// TIA Portal project "ModBus_Tcp_ESP32_V20" (V20)
// Modbus TCP/IP connection with ESP32 microcontroller

(* hardware
DEVICE "S7-1200 station_1"  S7-1200 Station
   slot 0: "Rack_0"  S7-1200 Rack  Rack  V1.0
   slot 1: "PLC_1"  CPU 1212C AC/DC/Rly  6ES7 212-1BE40-0XB0  V4.6
DEVICE "HMI_1"  TP700 Comfort
   slot 0: "HMI_1"  TP700 Comfort  6AV2 124-0GC01-0AX0  17.0.0.0
   slot 1: "HMI_RT_1"  TP700 Comfort  6AV2 124-0GC01-0AX0  17.0.0.0
   slot 5: "HMI_1.IE_CP_1"  PROFINET Interface  17.0.0.0
      slot 1: "PROFINET Interface_1"  PROFINET Interface
         slot 1: "Port_1"  Port
         slot 2: "Port_2"  Port
   slot 7: "HMI_1.MPI/DP_CP_1"  MPI/DP Interface  17.0.0.0
*)

// ===== PLC "PLC_1"  CPU 1212C AC/DC/Rly =====

VAR_GLOBAL   // PLC tag table "Default tag table"
   "Clock_Byte" AT %MB0 : Byte;
   "Clock_10Hz" AT %M0.0 : Bool;
   "Clock_5Hz" AT %M0.1 : Bool;
   "Clock_2.5Hz" AT %M0.2 : Bool;
   "Clock_2Hz" AT %M0.3 : Bool;
   "Clock_1.25Hz" AT %M0.4 : Bool;
   "Clock_1Hz" AT %M0.5 : Bool;
   "Clock_0.625Hz" AT %M0.6 : Bool;
   "Clock_0.5Hz" AT %M0.7 : Bool;
   "Tag_1" AT %MW1 : Word;
   "Tag_2" AT %M10.1 : Bool;
   "Tag_3" AT %M10.5 : Bool;
   "Tag_4" AT %M100.1 : Bool;
   "Tag_5" AT %M10.6 : Bool;
   "Tag_6" AT %M11.1 : Bool;
   "Tag_7" AT %M12.1 : Bool;
   "Tag_8" AT %M10.0 : Bool;
END_VAR

DATA_BLOCK "Modbus_Receiver"   // DB2
{ S7_Optimized_Access := 'FALSE' }
VERSION : 0.1
   VAR
      Receiver : Array[0..7] of Word;
      ADDR : UDInt := 400001;   // Initial Address Holding Register
      DATA_LEN : UInt := 8;   // Holding Register to Read
   END_VAR
BEGIN
   // Receiver[0] : First Address
   // Receiver[4] : Command
   // Receiver[3] : Value
   // Receiver[2] : Third Address
   // Receiver[1] : Second Address
   // Receiver[5] : Frequency Readed
   // Receiver[6] : Output Current
   // Receiver[7] : Drive Status
END_DATA_BLOCK

DATA_BLOCK "Param_Modbus"   // DB3
{ S7_Optimized_Access := 'FALSE' }
VERSION : 0.1
   VAR
      Receiver : Struct
         Request : Bool := true;
         Error : Bool;
         Disconnect : Bool := false;
         NDR : Bool;
         DR : Bool;
         Status : Word;
         Done : Bool;
         Busy : Bool;
         Mb_Mode : Int := 0;
         Rev_Connection : TCON_IP_v4;
      END_STRUCT;
      Sender : Struct
         Request : Bool := true;
         Error : Bool;
         Disconnect : Bool;
         NDR : Bool;
         DR : Bool;
         Status : Word;
         Done : Bool;
         Busy : Bool;
         Mb_Mode : Int := 1;
         Sen_Connection : TCON_IP_v4;
      END_STRUCT;
   END_VAR
BEGIN
   Receiver.Rev_Connection.InterfaceId := 64;
   Receiver.Rev_Connection.ID := 1;
   Receiver.Rev_Connection.ConnectionType := 11;
   Receiver.Rev_Connection.ActiveEstablished := true;
   Receiver.Rev_Connection.RemoteAddress.ADDR[1] := 192;
   Receiver.Rev_Connection.RemoteAddress.ADDR[2] := 168;
   Receiver.Rev_Connection.RemoteAddress.ADDR[3] := 20;
   Receiver.Rev_Connection.RemoteAddress.ADDR[4] := 55;
   Receiver.Rev_Connection.RemotePort := 502;
   Receiver.Rev_Connection.LocalPort := 502;
   Sender.Sen_Connection.InterfaceId := 64;
   Sender.Sen_Connection.ID := 1;
   Sender.Sen_Connection.ConnectionType := 11;
   Sender.Sen_Connection.ActiveEstablished := true;
   Sender.Sen_Connection.RemoteAddress.ADDR[1] := 192;
   Sender.Sen_Connection.RemoteAddress.ADDR[2] := 168;
   Sender.Sen_Connection.RemoteAddress.ADDR[3] := 20;
   Sender.Sen_Connection.RemoteAddress.ADDR[4] := 55;
   Sender.Sen_Connection.RemotePort := 502;
   Sender.Sen_Connection.LocalPort := 502;
END_DATA_BLOCK

DATA_BLOCK "Modbus_Sender"   // DB5
{ S7_Optimized_Access := 'FALSE' }
VERSION : 0.1
   VAR
      Sending : Array[0..4] of Int;
      bitStartStop : Int;   // Bit de habilitar o deshabilitar variador
      ADDR : UDInt := 400001;   // Holding Register desde el cual iniciara a escribir
      DATA_LEN : UInt := 5;   // Numero de Holding Register de escritura
   END_VAR
BEGIN
   // Sending[0] : Address 1
   // Sending[1] : Address 2
   // Sending[2] : Address 3
   // Sending[3] : Value
   // Sending[4] : Command
END_DATA_BLOCK

DATA_BLOCK "DATA"   // DB9
{ S7_Optimized_Access := 'TRUE' }
VERSION : 0.1
   VAR
      HMI_DATA : Struct   // Vars for inputs and outputs displayed in HMI
         Inputs : Struct
            setFrequency : Bool;   // Setpoint frequency x10, e.g. 100 = 10.0Hz
            frequencySetPoint : Int;   // Write frequency value
            startVFD : Bool;   // Write 1 to address
            stopVFD : Bool;   // Write 0 to address
         END_STRUCT;
         Outputs : Struct
            outputFrequency : Int;   // Output frequency value
            outputCurrent : Int;   // Output current value
            driveStatus : Bool;   // 0 = Stop / 1 = Run Enable
         END_STRUCT;
      END_STRUCT;
      Connect_Disconnect : Struct   // Vars for disconnect MB_Client block
         bitVFD : Bool;
         setFrequency : Bool;
         driveStatus : Bool;
         outputCurrent : Bool;
         outputFrequency : Bool;
         disconnectMBWrite : Bool;
         disconnectMBRead : Bool;
         disconnectSignal : Bool;   // Disconnect signal for MB_Client
      END_STRUCT;
      bitStop : Bool;   // Feedback Stopt from HMI
      bitStart : Bool;   // Feedback Start from HMI
      counterValue : Int;   // Counter current value
      RisingEdgeCounter : Bool;   // Memory for rising edge for counter activate
      disableCounter : Bool;
   END_VAR
BEGIN
END_DATA_BLOCK

FUNCTION "Write_Data" : Void   // FC1, LAD
{ S7_Optimized_Access := 'TRUE' }
VERSION : 0.1
   VAR_TEMP   // added for the SCL form of the ladder/FBD networks
      _w1 : Bool;
   END_VAR
BEGIN

REGION Network 1: Start or Stop VFD
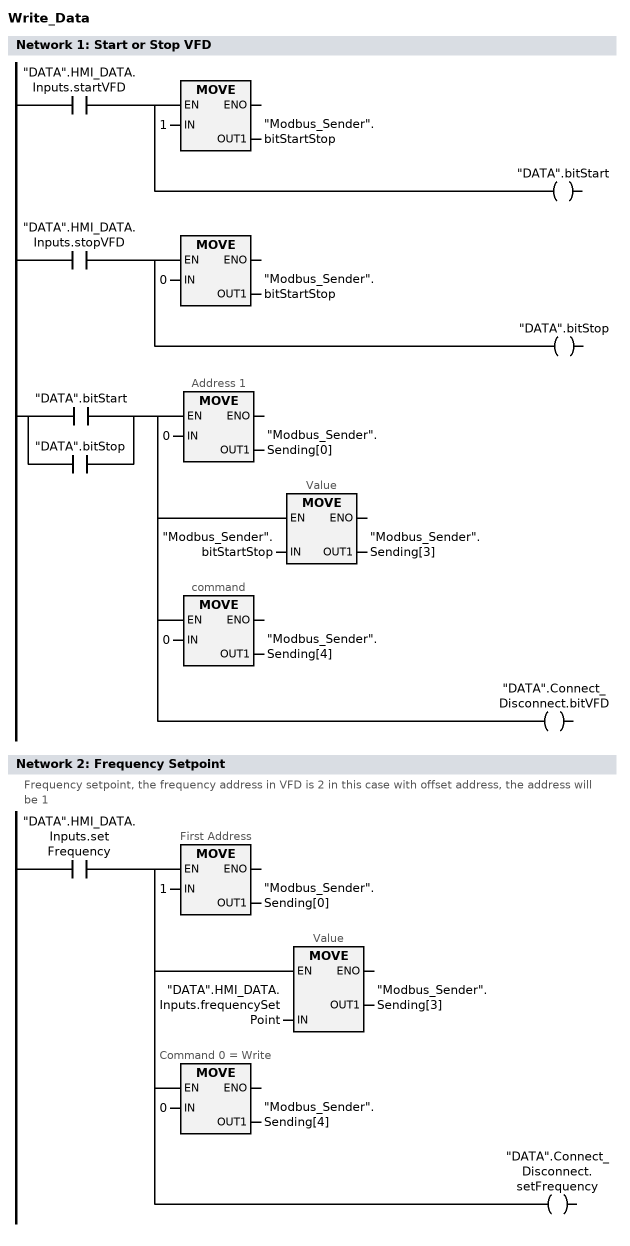
   RUNG wire#powerrail
      Contact( "DATA".HMI_DATA.Inputs.startVFD )
      wire#w1
      Move(in := 1, out1 => "Modbus_Sender".bitStartStop)
   END_RUNG
   RUNG wire#w1
      Coil( "DATA".bitStart )
   END_RUNG
   RUNG wire#powerrail
      Contact( "DATA".HMI_DATA.Inputs.stopVFD )
      wire#w2
      Move(in := 0, out1 => "Modbus_Sender".bitStartStop)
   END_RUNG
   RUNG wire#w2
      Coil( "DATA".bitStop )
   END_RUNG
   RUNG wire#powerrail
      Contact( "DATA".bitStart )
      wire#w3
      Move(in := 0, out1 => "Modbus_Sender".Sending[0])   // Address 1
   END_RUNG
   RUNG wire#powerrail
      Contact( "DATA".bitStop )
   END_RUNG wire#w3
   RUNG wire#w3
      Move(in := "Modbus_Sender".bitStartStop, out1 => "Modbus_Sender".Sending[3])   // Value
   END_RUNG
   RUNG wire#w3
      Move(in := 0, out1 => "Modbus_Sender".Sending[4])   // command
   END_RUNG
   RUNG wire#w3
      Coil( "DATA".Connect_Disconnect.bitVFD )
   END_RUNG
   // the same network as SCL:
   IF "DATA".HMI_DATA.Inputs.startVFD THEN "Modbus_Sender".bitStartStop := 1; END_IF;
   "DATA".bitStart := "DATA".HMI_DATA.Inputs.startVFD;
   IF "DATA".HMI_DATA.Inputs.stopVFD THEN "Modbus_Sender".bitStartStop := 0; END_IF;
   "DATA".bitStop := "DATA".HMI_DATA.Inputs.stopVFD;
   #_w1 := "DATA".bitStart OR "DATA".bitStop;
   IF #_w1 THEN
       "Modbus_Sender".Sending[0] := 0;   // Address 1
       "Modbus_Sender".Sending[3] := "Modbus_Sender".bitStartStop;   // Value
       "Modbus_Sender".Sending[4] := 0;   // command
   END_IF;
   "DATA".Connect_Disconnect.bitVFD := #_w1;
END_REGION

REGION Network 2: Frequency Setpoint
   // Frequency setpoint, the frequency address in VFD is 2 in this case with offset address, the address will be 1
   RUNG wire#powerrail
      Contact( "DATA".HMI_DATA.Inputs.setFrequency )
      wire#w1
      Move(in := 1, out1 => "Modbus_Sender".Sending[0])   // First Address
   END_RUNG
   RUNG wire#w1
      Move(in := "DATA".HMI_DATA.Inputs.frequencySetPoint, out1 => "Modbus_Sender".Sending[3])   // Value
   END_RUNG
   RUNG wire#w1
      Move(in := 0, out1 => "Modbus_Sender".Sending[4])   // Command 0 = Write
   END_RUNG
   RUNG wire#w1
      Coil( "DATA".Connect_Disconnect.setFrequency )
   END_RUNG
   // the same network as SCL:
   IF "DATA".HMI_DATA.Inputs.setFrequency THEN
       "Modbus_Sender".Sending[0] := 1;   // First Address
       "Modbus_Sender".Sending[3] := "DATA".HMI_DATA.Inputs.frequencySetPoint;   // Value
       "Modbus_Sender".Sending[4] := 0;   // Command 0 = Write
   END_IF;
   "DATA".Connect_Disconnect.setFrequency := "DATA".HMI_DATA.Inputs.setFrequency;
END_REGION
END_FUNCTION

FUNCTION "Read_Data" : Void   // FC2, LAD
TITLE = Read data from VFD, each modbus address have offset of 1. eg. for address 1 in VFD, the modbus address will be 0
{ S7_Optimized_Access := 'TRUE' }
VERSION : 0.1
   VAR_TEMP   // added for the SCL form of the ladder/FBD networks
      _w1 : Bool;
   END_VAR
BEGIN

REGION Network 1: Counter
   // Counter conditional for each read instruction
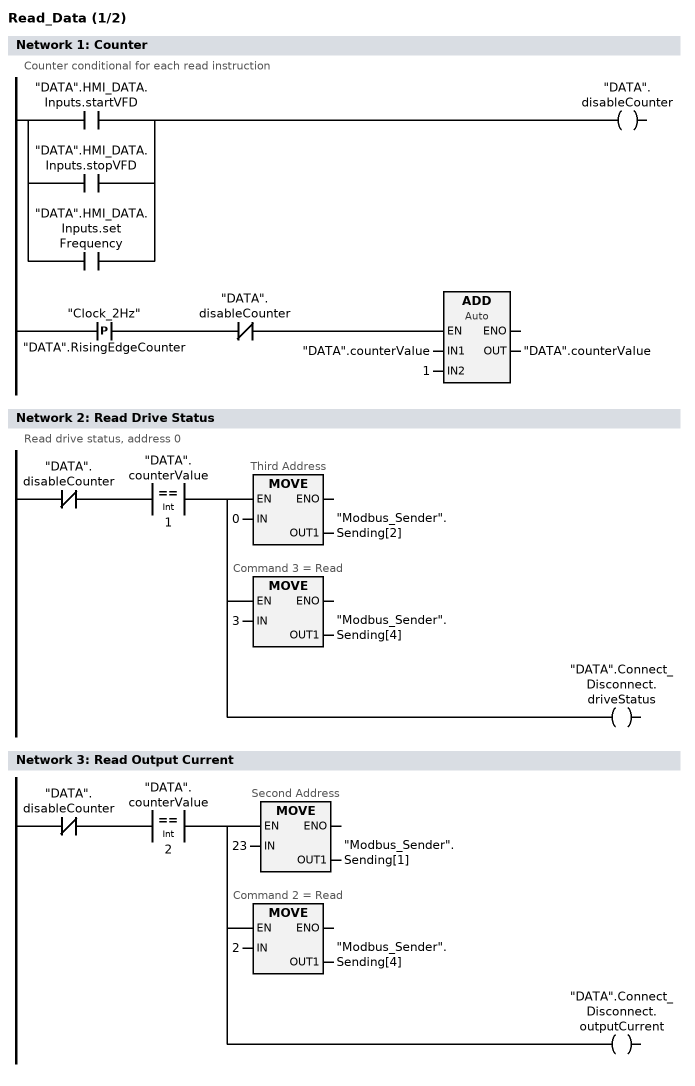
   RUNG wire#powerrail
      Contact( "DATA".HMI_DATA.Inputs.startVFD )
      wire#w1
      Coil( "DATA".disableCounter )
   END_RUNG
   RUNG wire#powerrail
      Contact( "DATA".HMI_DATA.Inputs.stopVFD )
   END_RUNG wire#w1
   RUNG wire#powerrail
      Contact( "DATA".HMI_DATA.Inputs.setFrequency )
   END_RUNG wire#w1
   RUNG wire#powerrail
      P_Contact(operand := "Clock_2Hz", bit := "DATA".RisingEdgeCounter)
      I_Contact( "DATA".disableCounter )
      Add(in1 := "DATA".counterValue, in2 := 1, out => "DATA".counterValue)
   END_RUNG
   // the same network as SCL:
   "DATA".disableCounter := "DATA".HMI_DATA.Inputs.startVFD OR "DATA".HMI_DATA.Inputs.stopVFD OR "DATA".HMI_DATA.Inputs.setFrequency;
   #_w1 := "Clock_2Hz" AND NOT "DATA".RisingEdgeCounter;   // rising edge of "Clock_2Hz"
   "DATA".RisingEdgeCounter := "Clock_2Hz";
   IF #_w1 AND NOT "DATA".disableCounter THEN "DATA".counterValue := "DATA".counterValue + 1; END_IF;
END_REGION

REGION Network 2: Read Drive Status
   // Read drive status, address 0
   RUNG wire#powerrail
      I_Contact( "DATA".disableCounter )
      { S7_Templates := "SrcType := Int" } EQ_Contact(in1 := "DATA".counterValue, in2 := 1)
      wire#w1
      Move(in := 0, out1 => "Modbus_Sender".Sending[2])   // Third Address
   END_RUNG
   RUNG wire#w1
      Move(in := 3, out1 => "Modbus_Sender".Sending[4])   // Command 3 = Read
   END_RUNG
   RUNG wire#w1
      Coil( "DATA".Connect_Disconnect.driveStatus )
   END_RUNG
   // the same network as SCL:
   #_w1 := NOT "DATA".disableCounter AND ("DATA".counterValue = 1);
   IF #_w1 THEN
       "Modbus_Sender".Sending[2] := 0;   // Third Address
       "Modbus_Sender".Sending[4] := 3;   // Command 3 = Read
   END_IF;
   "DATA".Connect_Disconnect.driveStatus := #_w1;
END_REGION

REGION Network 3: Read Output Current
   RUNG wire#powerrail
      I_Contact( "DATA".disableCounter )
      { S7_Templates := "SrcType := Int" } EQ_Contact(in1 := "DATA".counterValue, in2 := 2)
      wire#w1
      Move(in := 23, out1 => "Modbus_Sender".Sending[1])   // Second Address
   END_RUNG
   RUNG wire#w1
      Move(in := 2, out1 => "Modbus_Sender".Sending[4])   // Command 2 = Read
   END_RUNG
   RUNG wire#w1
      Coil( "DATA".Connect_Disconnect.outputCurrent )
   END_RUNG
   // the same network as SCL:
   #_w1 := NOT "DATA".disableCounter AND ("DATA".counterValue = 2);
   IF #_w1 THEN
       "Modbus_Sender".Sending[1] := 23;   // Second Address
       "Modbus_Sender".Sending[4] := 2;   // Command 2 = Read
   END_IF;
   "DATA".Connect_Disconnect.outputCurrent := #_w1;
END_REGION

REGION Network 4: Read Frequency
   // Lectura de valor de frecuencia, direccion con offset de 1
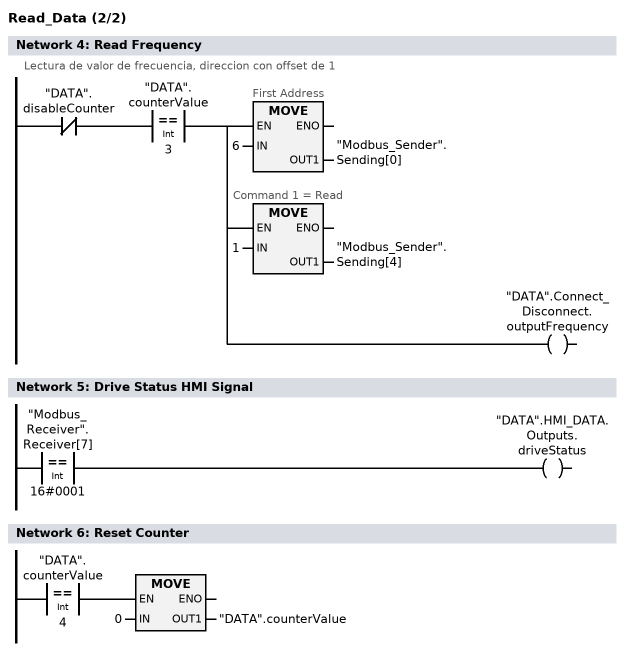
   RUNG wire#powerrail
      I_Contact( "DATA".disableCounter )
      { S7_Templates := "SrcType := Int" } EQ_Contact(in1 := "DATA".counterValue, in2 := 3)
      wire#w1
      Move(in := 6, out1 => "Modbus_Sender".Sending[0])   // First Address
   END_RUNG
   RUNG wire#w1
      Move(in := 1, out1 => "Modbus_Sender".Sending[4])   // Command 1 = Read
   END_RUNG
   RUNG wire#w1
      Coil( "DATA".Connect_Disconnect.outputFrequency )
   END_RUNG
   // the same network as SCL:
   #_w1 := NOT "DATA".disableCounter AND ("DATA".counterValue = 3);
   IF #_w1 THEN
       "Modbus_Sender".Sending[0] := 6;   // First Address
       "Modbus_Sender".Sending[4] := 1;   // Command 1 = Read
   END_IF;
   "DATA".Connect_Disconnect.outputFrequency := #_w1;
END_REGION

REGION Network 5: Drive Status HMI Signal
   RUNG wire#powerrail
      { S7_Templates := "SrcType := Int" } EQ_Contact(in1 := "Modbus_Receiver".Receiver[7], in2 := 16#0001)
      Coil( "DATA".HMI_DATA.Outputs.driveStatus )
   END_RUNG
   // the same network as SCL:
   "DATA".HMI_DATA.Outputs.driveStatus := "Modbus_Receiver".Receiver[7] = 16#0001;
END_REGION

REGION Network 6: Reset Counter
   RUNG wire#powerrail
      { S7_Templates := "SrcType := Int" } EQ_Contact(in1 := "DATA".counterValue, in2 := 4)
      Move(in := 0, out1 => "DATA".counterValue)
   END_RUNG
   // the same network as SCL:
   IF "DATA".counterValue = 4 THEN "DATA".counterValue := 0; END_IF;
END_REGION
END_FUNCTION

FUNCTION "MB_CLIENT_R/W" : Void   // FC3, LAD
{ S7_Optimized_Access := 'TRUE' }
VERSION : 0.1
BEGIN

REGION Network 1 (SCL): Disconnect signal for each MB_CLIENT block depending of the function to execute
   IF ("DATA".Connect_Disconnect.bitVFD OR "DATA".Connect_Disconnect.setFrequency OR "DATA".Connect_Disconnect.driveStatus OR "DATA".Connect_Disconnect.outputCurrent OR "DATA".Connect_Disconnect.outputFrequency) THEN
       "DATA".Connect_Disconnect.disconnectSignal := TRUE;
   ELSE
       "DATA".Connect_Disconnect.disconnectSignal := FALSE;
   END_IF;
END_REGION

REGION Network 2: Read ModbusRTU Data
   // Read ModbusRTU Data from drive via ModbusTCP/IP ESP32
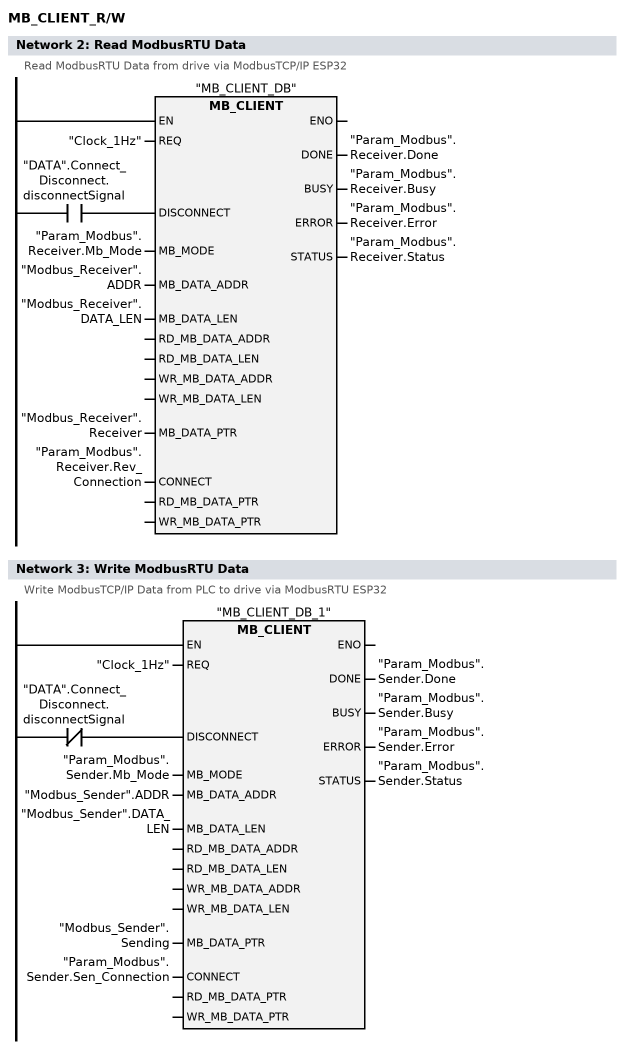
   "MB_CLIENT_DB"(REQ := "Clock_1Hz",   // MB_CLIENT
                  DISCONNECT := "DATA".Connect_Disconnect.disconnectSignal,
                  MB_MODE := "Param_Modbus".Receiver.Mb_Mode,
                  MB_DATA_ADDR := "Modbus_Receiver".ADDR,
                  MB_DATA_LEN := "Modbus_Receiver".DATA_LEN,
                  MB_DATA_PTR := "Modbus_Receiver".Receiver,
                  CONNECT := "Param_Modbus".Receiver.Rev_Connection,
                  DONE => "Param_Modbus".Receiver.Done,
                  BUSY => "Param_Modbus".Receiver.Busy,
                  ERROR => "Param_Modbus".Receiver.Error,
                  STATUS => "Param_Modbus".Receiver.Status);
END_REGION

REGION Network 3: Write ModbusRTU Data
   // Write ModbusTCP/IP Data from PLC to drive via ModbusRTU ESP32
   "MB_CLIENT_DB_1"(REQ := "Clock_1Hz",   // MB_CLIENT
                    DISCONNECT := NOT "DATA".Connect_Disconnect.disconnectSignal,
                    MB_MODE := "Param_Modbus".Sender.Mb_Mode,
                    MB_DATA_ADDR := "Modbus_Sender".ADDR,
                    MB_DATA_LEN := "Modbus_Sender".DATA_LEN,
                    MB_DATA_PTR := "Modbus_Sender".Sending,
                    CONNECT := "Param_Modbus".Sender.Sen_Connection,
                    DONE => "Param_Modbus".Sender.Done,
                    BUSY => "Param_Modbus".Sender.Busy,
                    ERROR => "Param_Modbus".Sender.Error,
                    STATUS => "Param_Modbus".Sender.Status);
END_REGION
END_FUNCTION

ORGANIZATION_BLOCK "Main"   // OB1, LAD, ProgramCycle
TITLE = "Main Program Sweep (Cycle)"
{ S7_Optimized_Access := 'TRUE' }
VERSION : 0.1
// Las direccion de registro tienen un offset de 1
// Las variables Disconnect de cada bloque modbus no pueden estar en FALSE al tiempo, por lo cual se realiza una logica con contactos para que cuando se este escribiendo, la variable disconnect del bloque de lectura este en TRUE y viceversa.
   VAR_INPUT
      Initial_Call : Bool;   // Initial call of this OB
      Remanence : Bool;   // =True, if remanent data are available
   END_VAR
BEGIN

REGION Network 1
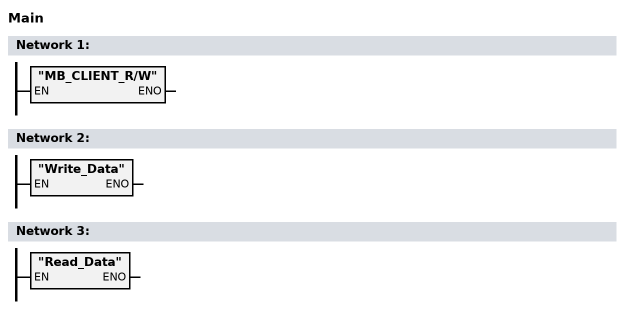
   RUNG wire#powerrail
      "MB_CLIENT_R/W"()
   END_RUNG
   // the same network as SCL:
   "MB_CLIENT_R/W"();
END_REGION

REGION Network 2
   RUNG wire#powerrail
      "Write_Data"()
   END_RUNG
   // the same network as SCL:
   "Write_Data"();
END_REGION

REGION Network 3
   RUNG wire#powerrail
      "Read_Data"()
   END_RUNG
   // the same network as SCL:
   "Read_Data"();
END_REGION
END_ORGANIZATION_BLOCK

(* ===== HMI "HMI_RT_1" =====
system functions are stored by id; their names below are inferred from use
connection "HMI_Connection_1": ETHERNET, S7_1200_OMS

HMI tags "Default tag table"
   "Tag_ScreenNumber" : UInt, internal
   "driveStatus" : Bool = PLC DATA.HMI_DATA.Outputs.driveStatus AT %DB1.DBX0.0, 100 ms
   "outputFrequency" : Word = PLC Modbus_Receiver.Receiver[5] AT %DB2.DBW10, 100 ms
   "outputCurrent" : Word = PLC Modbus_Receiver.Receiver[6] AT %DB2.DBW12, 100 ms
   "frequencySetPoint" : Int = PLC DATA.HMI_DATA.Inputs.frequencySetPoint AT %DB1.DBW0, 1 s
   "setFrequency" : Bool = PLC DATA.HMI_DATA.Inputs.setFrequency AT %DB1.DBX0.0, 1 s
   "startVFD" : Bool = PLC DATA.HMI_DATA.Inputs.startVFD AT %DB1.DBX0.0, 1 s
   "stopVFD" : Bool = PLC DATA.HMI_DATA.Inputs.stopVFD AT %DB1.DBX0.0, 1 s

screen "Root screen" 800x420, template "Template_1"
   on GenerateScreen: SetTag("Tag_ScreenNumber", 1)
   GraphicView "Graphic view_1" at 309,13 size 187x105; Picture "Graphic_5"
   GraphicView "Graphic view_2" at 309,13 size 187x105; Picture "Graphic_7"
      Visibility <- "driveStatus"
   IOField "I/O field_1" at 240,153 size 92x39; FormatPattern 9999
      ProcessValue <- "outputFrequency"
   IOField "I/O field_2" at 474,154 size 73x38; FormatPattern 999
      ProcessValue <- "outputCurrent"
   TextField "Text field_1" at 240,123 size 97x23; Text 'Frequency'
   TextField "Text field_2" at 440,123 size 142x23; Text 'Output Current'
   Button "Button_1" at 115,237 size 96x32; TextOff 'Start VFD'
      on Press: function_b14e0dd5("startVFD", 0)
   Button "Button_2" at 115,283 size 96x32; TextOff 'Stop VFD'
      on Press: function_b14e0dd5("stopVFD", 0)
   IOField "I/O field_3" at 462,277 size 96x32; FormatPattern 999
      ProcessValue <- "frequencySetPoint"
   TextField "Text field_3" at 435,246 size 180x23; Text 'Frequency Setpoint'
   Button "Button_3" at 578,277 size 96x32; TextOff 'Set Hz'
      on Press: function_b14e0dd5("setFrequency", 0)

Template "Template_1" 800x420
   Button "Exit" at 720,360 size 78x58; TextOff 'Exit'; PictureOff "ExitRuntime_TP700_Comfort_TR"; PictureOn "ExitRuntime_TP700_Comfort_TR"
      on Release: StopRuntime(0)
   Button "Template_Button" at 640,360 size 78x58; TextOff 'Text'
   Button "Template_Button_1" at 560,360 size 78x58; TextOff 'Text'
   Button "Template_Button_2" at 480,360 size 78x58; TextOff 'Text'
   Button "Template_Button_3" at 400,360 size 78x58; TextOff 'Text'
   Button "Template_Button_4" at 321,360 size 78x58; TextOff 'Text'
   Button "Template_Button_5" at 241,360 size 78x58; TextOff 'Text'
   Button "Template_Button_6" at 161,360 size 78x58; TextOff 'Text'
   Button "Template_Button_7" at 81,360 size 78x58; TextOff 'Text'
   Button "Start screen" at 1,360 size 78x58; TextOff 'Start screen'; PictureOff "NavigateHome_TP700_Comfort_TR"; PictureOn "NavigateHome_TP700_Comfort_TR"
      on Release: ActivateScreen("Root screen", 0)
*)